screen "10_Startscreen" 800x480, template "01_Navigation"
   on GenerateScreen: SetTag("MainNavigationState", 1)
   GraphicView "Graphic view_2" at 0,0 size 800x480; Picture "PopUpBackground"
      Visibility <- "PopUpBackground"
   Button "Button_7" at 14,136 size 30x30; TextOff 'Text'
      Visibility <- "DB_HMI_Global_selection"
   Button "Button_10" at 14,195 size 30x30; TextOff 'Text'
      Visibility <- "DB_HMI_Global_selection"
   Button "Button_11" at 14,250 size 30x30; TextOff 'Text'
      Visibility <- "DB_HMI_Global_selection"
   Button "Button_13" at 14,311 size 30x30; TextOff 'Text'
      Visibility <- "DB_HMI_Global_selection"
   TextField "txtContentboard1" at 667,136 size 59x34; Text 'Calc. Time [s] / Name Parameter'
   TextField "txtContentboard1_1" at 723,141 size 65x24; Text 'Meas. Time [s] / Name Parameter'
   Button "Button_1" at 14,136 size 30x30; TextOff 'Text'
      on Click: SetTag("DB_HMI_Global_selection", 3)
   Button "Button_2" at 14,195 size 30x30; TextOff 'Text'
      on Click: SetTag("DB_HMI_Global_selection", 4)
   Button "Button_3" at 14,251 size 30x30; TextOff 'Text'
      on Click: SetTag("DB_HMI_Global_selection", 6)
   Button "Button_12" at 14,310 size 30x30; TextOff 'Text'
      on Click: SetTag("DB_HMI_Global_selection", 0)
   TextField "txtParameter1" at 82,159 size 99x24; Text 'Status / Parameter 1'
      Visibility <- "InScreenTabState"
   TextField "txtParameter1_1" at 82,199 size 99x24; Text 'Mode / Parameter 1'
      Visibility <- "InScreenTabState"
   TextField "txtParameter1_3" at 83,242 size 84x24; Text 'Producing car / Parameter 1'
      Visibility <- "InScreenTabState"
   TextField "Text field_4" at 32,381 size 142x20; Text 'Operation Commands'
   TextField "Text field_1" at 32,99 size 105x20; Text 'Production Line'
   TextField "txtParameter1_2" at 194,159 size 99x24; Text 'Status / Parameter 1'
      Visibility <- "InScreenTabState"
   TextField "txtParameter1_4" at 195,197 size 99x24; Text 'Mode / Parameter 1'
      Visibility <- "InScreenTabState"
   TextField "txtParameter1_5" at 195,242 size 84x24; Text 'Producing car / Parameter 1'
      Visibility <- "InScreenTabState"
   TextField "txtParameter1_6" at 306,159 size 99x24; Text 'Status / Parameter 1'
      Visibility <- "InScreenTabState"
   TextField "txtParameter1_7" at 307,197 size 99x24; Text 'Mode / Parameter 1'
      Visibility <- "InScreenTabState"
   TextField "txtParameter1_8" at 307,242 size 84x24; Text 'Producing car / Parameter 1'
      Visibility <- "InScreenTabState"
   TextField "txtParameter1_9" at 418,159 size 99x24; Text 'Status / Parameter 1'
      Visibility <- "InScreenTabState"
   TextField "txtParameter1_10" at 419,197 size 99x24; Text 'Mode / Parameter 1'
      Visibility <- "InScreenTabState"
   TextField "txtParameter1_11" at 419,242 size 84x24; Text 'Producing car / Parameter 1'
      Visibility <- "InScreenTabState"
   TextField "txtParameter1_12" at 530,159 size 99x24; Text 'Status / Parameter 1'
      Visibility <- "InScreenTabState"
   TextField "txtParameter1_13" at 531,197 size 99x24; Text 'Mode / Parameter 1'
      Visibility <- "InScreenTabState"
   TextField "txtParameter1_14" at 531,242 size 84x24; Text 'Producing car / Parameter 1'
      Visibility <- "InScreenTabState"
   GraphicView "Graphic view_1" at 46,139 size 25x25; Picture "Car_Red"
   GraphicView "Graphic view_3" at 47,196 size 25x25; Picture "Car_Green"
   GraphicView "Graphic view_4" at 47,251 size 25x25; Picture "Car_Blue_1"
   IOField "I/O field_1" at 671,168 size 56x24; FormatPattern 999
      ProcessValue <- "DB_HMI_ARG1_Seq1_Calculated_PT_Red(4)"
   TextField "txtTitleBar" at 80,128 size 55x24; Text 'Station 1 / Applikation'
   GraphicView "Graphic view_5" at 636,169 size 25x25; Picture "Car_Red"
   GraphicView "Graphic view_6" at 636,226 size 25x25; Picture "Car_Green"
   GraphicView "Graphic view_7" at 636,285 size 25x25; Picture "Car_Blue_1"
   TextField "txtTitleBar_1" at 200,122 size 55x24; Text 'Station 2 / Applikation'
   TextField "txtTitleBar_2" at 320,122 size 55x24; Text 'Station 3 / Applikation'
   TextField "txtTitleBar_3" at 440,122 size 55x24; Text 'Station 4 / Applikation'
   TextField "txtTitleBar_4" at 560,122 size 55x24; Text 'Station 5 / Applikation'
   Button "btnStart" at 184,377 size 119x29; TextOn 'STOP'; TextOff 'START'
      on Press: SetTag("DB_HMI_Global_Cmd_Start", 1); SetTag("DB_HMI_Global_Cmd_Start(1)", 1); SetTag("DB_HMI_Global_Cmd_Start(2)", 1); SetTag("DB_HMI_Global_Cmd_Start(3)", 1); SetTag("DB_HMI_Global_Cmd_Start(4)", 1)
      on Release: SetTag("DB_HMI_Global_Cmd_Start", 0); SetTag("DB_HMI_Global_Cmd_Start(1)", 0); SetTag("DB_HMI_Global_Cmd_Start(2)", 0); SetTag("DB_HMI_Global_Cmd_Start(3)", 0); SetTag("DB_HMI_Global_Cmd_Start(4)", 0)
   Button "btnStart_1" at 312,376 size 120x30; TextOn 'STOP'; TextOff 'STOP / START'
      on Release: SetTag("DB_HMI_Global_Cmd_Stop", 0); SetTag("DB_HMI_Global_Cmd_Stop(1)", 0); SetTag("DB_HMI_Global_Cmd_Stop(2)", 0); SetTag("DB_HMI_Global_Cmd_Stop(3)", 0); SetTag("DB_HMI_Global_Cmd_Stop(4)", 0)
      on Press: SetTag("DB_HMI_Global_Cmd_Stop", 1); SetTag("DB_HMI_Global_Cmd_Stop(1)", 1); SetTag("DB_HMI_Global_Cmd_Stop(2)", 1); SetTag("DB_HMI_Global_Cmd_Stop(3)", 1); SetTag("DB_HMI_Global_Cmd_Stop(4)", 1)
   IOField "I/O field_2" at 727,168 size 56x24; FormatPattern 999
      ProcessValue <- "DB_HMI_ARG1_Seq1_Messured_PT_Red(4)"
   TextField "txtTitleBar_5" at 192,128 size 55x24; Text 'Station 2 / Applikation'
   TextField "txtTitleBar_6" at 304,128 size 55x24; Text 'Station 3 / Applikation'
   TextField "txtTitleBar_7" at 416,128 size 55x24; Text 'Station 4 / Applikation'
   TextField "Text field_52" at 81,297 size 549x14; Text 'Text'
   TextField "txtTitleBar_8" at 528,128 size 55x24; Text 'Station 5 / Applikation'
   IOField "I/O field_3" at 671,224 size 56x24; FormatPattern 999
      ProcessValue <- "DB_HMI_ARG1_Seq1_Calculated_PT_Green(4)"
   IOField "I/O field_4" at 727,224 size 56x24; FormatPattern 999
      ProcessValue <- "DB_HMI_ARG1_Seq1_Messured_PT_Green(4)"
   IOField "I/O field_5" at 671,280 size 56x24; FormatPattern 999
      ProcessValue <- "DB_HMI_ARG1_Seq1_Calculated_PT_Blue(4)"
   IOField "I/O field_6" at 727,280 size 56x24; FormatPattern 999
      ProcessValue <- "DB_HMI_ARG1_Seq1_Messured_PT_Blue(4)"
   GraphicView "Grafikanzeige_1" at 46,312 size 26x22; Picture "Grafik_4"
   Button "btnState" at 143,133 size 39x25; TextOff '...'; PictureOff "More_Icon"
      on Click: ActivateScreen("21_Station_1", 0); SetTag("SubNavigationState", 2)
   Button "btnState_1" at 255,133 size 39x25; TextOff '...'; PictureOff "More_Icon"
      on Click: ActivateScreen("22_Station_2", 0); SetTag("SubNavigationState", 3)
   Button "btnState_2" at 367,133 size 39x25; TextOff '...'; PictureOff "More_Icon"
      on Click: ActivateScreen("23_Station_3", 0); SetTag("SubNavigationState", 4)
   Button "btnState_3" at 479,133 size 39x25; TextOff '...'; PictureOff "More_Icon"
      on Click: ActivateScreen("24_Station_4", 0); SetTag("SubNavigationState", 5)
   Button "btnState_4" at 591,133 size 39x25; TextOff '...'; PictureOff "More_Icon"
      on Click: ActivateScreen("25_Station_5", 0); SetTag("SubNavigationState", 6)
   Rectangle "rectState" at 0,48 size 56x38
      Appearance <- "CurrentMachineState"
   Button "btnState_5" at 201,53 size 34x31; TextOff '...'; PictureOff "More_Icon"
      on Click: ActivateScreen("11_Mode_Global", 0)
   TextField "Auto" at 67,63 size 35x20; Text 'Auto'
      Visibility <- "DB_HMI_Global_Status_Auto"
   TextField "Manual" at 69,63 size 34x20; Text 'Man'
      Visibility <- "DB_HMI_Global_Status_Man"
   TextField "txtStateHeadline" at 65,48 size 123x23; Text 'Mode / Status'
   Button "sTATUS" at 80,184 size 102x25; TextOff 'Text'; TextList "MachineStatus"
      on Activate: "VBFunction_1"()
      ProcessValue <- "status"
   Button "sTATUS_1" at 192,184 size 102x25; TextOff 'Text'; TextList "MachineStatus"
      ProcessValue <- "DB_HMI_ARG1_Seq1_Status_Busy(1)"
   Button "sTATUS_2" at 304,184 size 102x25; TextOff 'Text'; TextList "MachineStatus"
      ProcessValue <- "DB_HMI_ARG1_Seq1_Status_Busy(2)"
   Button "sTATUS_3" at 416,184 size 102x25; TextOff 'Text'; TextList "MachineStatus"
      ProcessValue <- "DB_HMI_ARG1_Seq1_Status_Busy(3)"
   Button "sTATUS_4" at 528,184 size 102x25; TextOff 'Text'; TextList "MachineStatus"
      ProcessValue <- "DB_HMI_ARG1_Seq1_Status_Busy(4)"
   Button "sTATUS_5" at 82,214 size 102x25; TextOff 'Text'; TextList "MachineMode"
      ProcessValue <- "DB_HMI_ARG1_Seq1_Status_Auto"
   Button "sTATUS_6" at 192,214 size 102x25; TextOff 'Text'; TextList "MachineMode"
      ProcessValue <- "DB_HMI_ARG1_Seq1_Status_Auto(1)"
   Button "sTATUS_7" at 304,214 size 102x25; TextOff 'Text'; TextList "MachineMode"
      ProcessValue <- "DB_HMI_ARG1_Seq1_Status_Auto(2)"
   Button "sTATUS_8" at 416,214 size 102x25; TextOff 'Text'; TextList "MachineMode"
      ProcessValue <- "DB_HMI_ARG1_Seq1_Status_Auto(3)"
   Button "sTATUS_9" at 528,214 size 102x25; TextOff 'Text'; TextList "MachineMode"
      ProcessValue <- "DB_HMI_ARG1_Seq1_Status_Auto(4)"
   Button "Button_4" at 101,274 size 60x60; TextOff 'Text'; PictureList "CarColorsGraph"
      ProcessValue <- "DB_HMI_inProduction"
   Button "Button_5" at 214,274 size 60x60; TextOff 'Text'; PictureList "CarColorsGraph"
      ProcessValue <- "DB_HMI_inProduction(1)"
   Button "Button_6" at 327,274 size 60x60; TextOff 'Text'; PictureList "CarColorsGraph"
      ProcessValue <- "DB_HMI_inProduction(2)"
   Button "Button_8" at 439,274 size 60x60; TextOff 'Text'; PictureList "CarColorsGraph"
      ProcessValue <- "DB_HMI_inProduction(3)"
   Button "Button_9" at 550,274 size 60x60; TextOff 'Text'; PictureList "CarColorsGraph"
      ProcessValue <- "DB_HMI_inProduction(4)"

screen "11_Mode_Global" 800x480
   Button "Button_5" at 299,208 size 88x48; TextOff 'Stop / AUTO'
      on Press: SetTag("DB_HMI_Global_Cmd_Auto", 1); SetTag("DB_HMI_Global_Cmd_Auto(1)", 1); SetTag("DB_HMI_Global_Cmd_Auto(2)", 1); SetTag("DB_HMI_Global_Cmd_Auto(3)", 1); SetTag("DB_HMI_Global_Cmd_Auto(4)", 1)
      on Release: SetTag("DB_HMI_Global_Cmd_Auto", 0); SetTag("DB_HMI_Global_Cmd_Auto(1)", 0); SetTag("DB_HMI_Global_Cmd_Auto(2)", 0); SetTag("DB_HMI_Global_Cmd_Auto(3)", 0); SetTag("DB_HMI_Global_Cmd_Auto(4)", 0)
   Button "Button_6" at 405,208 size 88x48; TextOff 'Reset / MAN'
      on Press: SetTag("DB_HMI_Global_Cmd_Man", 1); SetTag("DB_HMI_Global_Cmd_Man(1)", 1); SetTag("DB_HMI_Global_Cmd_Man(2)", 1); SetTag("DB_HMI_Global_Cmd_Man(3)", 1); SetTag("DB_HMI_Global_Cmd_Man(4)", 1)
      on Release: SetTag("DB_HMI_Global_Cmd_Man", 0); SetTag("DB_HMI_Global_Cmd_Man(1)", 0); SetTag("DB_HMI_Global_Cmd_Man(2)", 0); SetTag("DB_HMI_Global_Cmd_Man(3)", 0); SetTag("DB_HMI_Global_Cmd_Man(4)", 0)
   Button "Button_1" at 177,283 size 440x40; TextOn 'CLOSE / SCHLIESSEN'; TextOff 'CLOSE / SCHLIESSEN'
      on Click: function_efd93a16()
      Appearance <- "ButtonDown"
   TextField "txtTitleBar" at 16,8 size 495x32; Text 'Operating Mode / Betriebsmodus'
   TextField "txtParameter7_3" at 193,122 size 163x24; Text 'Current Mode / Aktueller Modus'
   TextField "Manual" at 193,148 size 35x20; Text 'Man'
      Visibility <- "DB_HMI_Global_Status_Man"
   TextField "Auto" at 193,149 size 41x20; Text 'Auto'
      Visibility <- "DB_HMI_Global_Status_Auto"

screen "21_Station_1" 800x480, template "01_Navigation"
   Button "Button_11" at 24,220 size 272x40; TextOff 'Simulate Values / Alle Quittieren'; PictureOff "More_Icon"
      on ReleaseLeft: ResetBit("Ext_AckSafety_DB_ack")
      on PressLeft: SetBit("Ext_AckSafety_DB_ack")
      on Click: ActivateScreen("40_SimValues_1", 0)
      on Press: ActivateScreen("40_SimValues_1", 0)
   Button "Button_1" at 24,324 size 272x40; TextOff 'Start / Alle Quittieren'; PictureOff "More_Icon"
      on Release: SetTag("DB_HMI_ARG1_Seq1_Cmd_Start", 0)
      on PressLeft: SetBit("Ext_AckSafety_DB_ack")
      on ReleaseLeft: ResetBit("Ext_AckSafety_DB_ack")
      on Press: SetTag("DB_HMI_ARG1_Seq1_Cmd_Start", 1); SetTag("DB_HMI_ARG1_Seq1_Cmd_Stop", 0)
      Visibility <- "DB_HMI_ARG1_Seq1_Status_Man"
      ObjectEnable <- "DB_HMI_ARG1_Seq1_Cmd_Start"
   Button "Button_2" at 24,376 size 272x40; TextOff 'Stop + Reset / Alle Quittieren'; PictureOff "More_Icon"
      on Release: SetTag("DB_HMI_ARG1_Seq1_Cmd_Stop", 0)
      on PressLeft: SetBit("Ext_AckSafety_DB_ack")
      on ReleaseLeft: ResetBit("Ext_AckSafety_DB_ack")
      on Press: SetTag("DB_HMI_ARG1_Seq1_Cmd_Stop", 1); SetTag("DB_HMI_ARG1_Seq1_Cmd_Start", 0)
      Visibility <- "DB_HMI_ARG1_Seq1_Status_Man"
      ObjectEnable <- "DB_HMI_ARG1_Seq1_Cmd_Stop"
   TextField "Text field_1" at 16,192 size 166x25; Text 'Simulation timers'
   TextField "Text field_2" at 16,296 size 105x25; Text 'Commands'
   TextField "Text field_26" at 564,176 size 204x24; Text 'Branch2'
   TextField "Text field_3" at 16,104 size 61x25; Text 'Status'
   TextField "Text field_16" at 344,176 size 204x24; Text 'Branch1'
   TextField "Text field_17" at 344,104 size 230x25; Text 'Running step sequences'
   Button "Button_3" at 218,123 size 45x45; TextOff 'Text'; PictureList "CarColorsGraph"
      Visibility <- "DB_HMI_ARG1_Seq1_Status_Auto"
      ProcessValue <- "DB_HMI_inProduction"
   TextField "Text field_4" at 180,104 size 118x27; Text 'Produced car'
   TextField "Text field_7" at 344,200 size 204x24; Text 'Step 1'
   TextField "Text field_5" at 344,224 size 204x24; Text 'Step 2'
   TextField "Text field_6" at 344,248 size 204x24; Text 'Step 3'
   TextField "Text field_8" at 344,272 size 204x24; Text 'Step 4'
   TextField "Text field_9" at 344,296 size 204x24; Text 'Step 5'
   TextField "Text field_10" at 344,320 size 204x24; Text 'Step 6'
   TextField "Text field_11" at 344,344 size 204x24; Text 'Step 7'
   TextField "Text field_12" at 344,368 size 204x24; Text 'Step 8'
   TextField "Text field_15" at 564,200 size 204x24; Text 'Step 1'
   TextField "Text field_18" at 564,224 size 204x24; Text 'Step 2'
   TextField "Text field_19" at 564,248 size 204x24; Text 'Step 3'
   TextField "Text field_20" at 564,272 size 204x24; Text 'Step 4'
   TextField "Text field_21" at 564,296 size 204x24; Text 'Step 5'
   TextField "Text field_22" at 564,320 size 204x24; Text 'Step 6'
   TextField "Text field_23" at 564,344 size 204x24; Text 'Step 7'
   TextField "Text field_24" at 564,368 size 204x24; Text 'Step 8'
   TextField "Text field_25" at 564,392 size 204x24; Text 'Step 9'
   TextField "Text field_13" at 344,392 size 204x24; Text 'Step 9'
   TextField "Text field_14" at 344,138 size 204x24; Text 'Step 0'
   TextField "Text field_52" at 344,200 size 204x24; Text 'Step 1'
      Visibility <- "DB_HMI_ARG1_Seq1_S2"
   TextField "Text field_27" at 344,224 size 204x24; Text 'Step 2'
      Visibility <- "DB_HMI_ARG1_Seq1_S3"
   TextField "Text field_28" at 344,249 size 204x24; Text 'Step 3'
      Visibility <- "DB_HMI_ARG1_Seq1_S4"
   TextField "Text field_29" at 344,272 size 204x24; Text 'Step 4'
      Visibility <- "DB_HMI_ARG1_Seq1_S5"
   TextField "Text field_30" at 344,296 size 204x24; Text 'Step 5'
      Visibility <- "DB_HMI_ARG1_Seq1_S6"
   TextField "Text field_31" at 344,320 size 204x24; Text 'Step 6'
      Visibility <- "DB_HMI_ARG1_Seq1_S7"
   TextField "Text field_32" at 344,344 size 204x24; Text 'Step 7'
      Visibility <- "DB_HMI_ARG1_Seq1_S8"
   TextField "Text field_33" at 344,368 size 204x24; Text 'Step 8'
      Visibility <- "DB_HMI_ARG1_Seq1_S9"
   TextField "Text field_34" at 344,392 size 204x24; Text 'Step 9'
      Visibility <- "DB_HMI_ARG1_Seq1_S10"
   TextField "Text field_35" at 564,200 size 204x24; Text 'Step 1'
      Visibility <- "DB_HMI_ARG1_Seq1_S11"
   TextField "Text field_36" at 564,224 size 204x24; Text 'Step 2'
      Visibility <- "DB_HMI_ARG1_Seq1_S12"
   TextField "Text field_37" at 564,248 size 204x24; Text 'Step 3'
      Visibility <- "DB_HMI_ARG1_Seq1_S13"
   TextField "Text field_38" at 564,272 size 204x24; Text 'Step 4'
      Visibility <- "DB_HMI_ARG1_Seq1_S14"
   TextField "Text field_39" at 564,296 size 204x24; Text 'Step 5'
      Visibility <- "DB_HMI_ARG1_Seq1_S15"
   TextField "Text field_40" at 564,320 size 204x24; Text 'Step 6'
      Visibility <- "DB_HMI_ARG1_Seq1_S16"
   TextField "Text field_41" at 564,344 size 204x24; Text 'Step 7'
      Visibility <- "DB_HMI_ARG1_Seq1_S17"
   TextField "Text field_42" at 564,368 size 204x24; Text 'Step 8'
      Visibility <- "DB_HMI_ARG1_Seq1_S18"
   TextField "Text field_43" at 564,392 size 204x24; Text 'Step 9'
      Visibility <- "DB_HMI_ARG1_Seq1_S19"
   TextField "Text field_44" at 344,138 size 204x24; Text 'Step 0'
      Visibility <- "DB_HMI_ARG1_Seq1_S1"
   SymbolicIOField "Symbolic I/O field_1" at 182,129 size 117x32; TextOn '1'; TextOff '0'; TextList "Car_color"
      ProcessValue <- "DB_HMI_dropdown_selection"
      Visibility <- "DB_HMI_ARG1_Seq1_Status_Man"
   TextField "Busy" at 14,134 size 41x22; Text 'Busy'
      Visibility <- "DB_HMI_ARG1_Seq1_Status_Busy"
   TextField "Idle" at 14,134 size 35x22; Text 'Idle'
      Visibility <- "DB_HMI_ARG1_Seq1_Status_Idle"
   Rectangle "rectState" at 0,48 size 56x38
      Appearance <- "CurrentMachineState"
   Button "btnState" at 201,53 size 34x31; TextOff '...'; PictureOff "More_Icon"
      on Click: ActivateScreen("31_Mode_Station_1", 0)
   TextField "Auto" at 67,63 size 35x20; Text 'Auto'
      Visibility <- "DB_HMI_ARG1_Seq1_Status_Auto"
   TextField "Manual" at 69,63 size 34x20; Text 'Man'
      Visibility <- "DB_HMI_ARG1_Seq1_Status_Man"
   TextField "txtStateHeadline" at 65,48 size 123x23; Text 'Mode / Status'

screen "22_Station_2" 800x480, template "01_Navigation"
   Button "Button_11" at 24,220 size 272x40; TextOff 'Simulate Values / Alle Quittieren'; PictureOff "More_Icon"
      on ReleaseLeft: ResetBit("Ext_AckSafety_DB_ack")
      on PressLeft: SetBit("Ext_AckSafety_DB_ack")
      on Click: ActivateScreen("40_SimValues_2", 0)
   Button "Button_1" at 24,324 size 272x40; TextOff 'Start / Alle Quittieren'; PictureOff "More_Icon"
      on Release: SetTag("DB_HMI_ARG1_Seq1_Cmd_Start(1)", 0)
      on PressLeft: SetBit("Ext_AckSafety_DB_ack")
      on ReleaseLeft: ResetBit("Ext_AckSafety_DB_ack")
      on Press: SetTag("DB_HMI_ARG1_Seq1_Cmd_Start(1)", 1); SetTag("DB_HMI_ARG1_Seq1_Cmd_Stop(1)", 0)
      Visibility <- "DB_HMI_ARG1_Seq1_Status_Man(1)"
      ObjectEnable <- "DB_HMI_ARG1_Seq1_Cmd_Start(1)"
   Button "Button_2" at 24,376 size 272x40; TextOff 'Stop + Reset / Alle Quittieren'; PictureOff "More_Icon"
      on Release: SetTag("DB_HMI_ARG1_Seq1_Cmd_Stop(1)", 0)
      on PressLeft: SetBit("Ext_AckSafety_DB_ack")
      on ReleaseLeft: ResetBit("Ext_AckSafety_DB_ack")
      on Press: SetTag("DB_HMI_ARG1_Seq1_Cmd_Stop(1)", 1); SetTag("DB_HMI_ARG1_Seq1_Cmd_Start(1)", 0)
      Visibility <- "DB_HMI_ARG1_Seq1_Status_Man(1)"
      ObjectEnable <- "DB_HMI_ARG1_Seq1_Cmd_Stop(1)"
   TextField "Text field_1" at 16,192 size 166x25; Text 'Simulation timers'
   TextField "Text field_2" at 16,296 size 105x25; Text 'Commands'
   TextField "Text field_26" at 564,176 size 204x24; Text 'Branch2'
   TextField "Text field_3" at 16,104 size 61x25; Text 'Status'
   TextField "Text field_16" at 344,176 size 204x24; Text 'Branch1'
   SymbolicIOField "DropDownCars" at 182,129 size 117x32; TextOn '1'; TextOff '0'; TextList "Car_color"
      ProcessValue <- "DB_HMI_dropdown_selection(1)"
      Visibility <- "DB_HMI_ARG1_Seq1_Status_Man(1)"
   TextField "Text field_17" at 344,104 size 230x25; Text 'Running step sequences'
   TextField "Text field_4" at 180,104 size 118x27; Text 'Produced car'
   Button "Button_3" at 218,123 size 45x45; TextOff 'Text'; PictureList "CarColorsGraph"
      Visibility <- "DB_HMI_ARG1_Seq1_Status_Auto(1)"
      ProcessValue <- "DB_HMI_inProduction(1)"
   TextField "Text field_7" at 344,200 size 204x24; Text 'Step 1'
   TextField "Text field_5" at 344,224 size 204x24; Text 'Step 2'
   TextField "Text field_6" at 344,248 size 204x24; Text 'Step 3'
   TextField "Text field_8" at 344,272 size 204x24; Text 'Step 4'
   TextField "Text field_9" at 344,296 size 204x24; Text 'Step 5'
   TextField "Text field_10" at 344,320 size 204x24; Text 'Step 6'
   TextField "Text field_11" at 344,344 size 204x24; Text 'Step 7'
   TextField "Text field_12" at 344,368 size 204x24; Text 'Step 8'
   TextField "Text field_15" at 564,200 size 204x24; Text 'Step 1'
   TextField "Text field_18" at 564,224 size 204x24; Text 'Step 2'
   TextField "Text field_19" at 564,248 size 204x24; Text 'Step 3'
   TextField "Text field_20" at 564,272 size 204x24; Text 'Step 4'
   TextField "Text field_21" at 564,296 size 204x24; Text 'Step 5'
   TextField "Text field_22" at 564,320 size 204x24; Text 'Step 6'
   TextField "Text field_23" at 564,344 size 204x24; Text 'Step 7'
   TextField "Text field_24" at 564,368 size 204x24; Text 'Step 8'
   TextField "Text field_25" at 564,392 size 204x24; Text 'Step 9'
   TextField "Text field_13" at 344,392 size 204x24; Text 'Step 9'
   TextField "Text field_14" at 344,138 size 204x24; Text 'Step 0'
   TextField "Text field_52" at 344,200 size 204x24; Text 'Step 1'
      Visibility <- "DB_HMI_ARG1_Seq1_S2(1)"
   TextField "Text field_27" at 344,224 size 204x24; Text 'Step 2'
      Visibility <- "DB_HMI_ARG1_Seq1_S3(1)"
   TextField "Text field_28" at 344,249 size 204x24; Text 'Step 3'
      Visibility <- "DB_HMI_ARG1_Seq1_S4(1)"
   TextField "Text field_29" at 344,272 size 204x24; Text 'Step 4'
      Visibility <- "DB_HMI_ARG1_Seq1_S5(1)"
   TextField "Text field_30" at 344,296 size 204x24; Text 'Step 5'
      Visibility <- "DB_HMI_ARG1_Seq1_S6(1)"
   TextField "Text field_31" at 344,320 size 204x24; Text 'Step 6'
      Visibility <- "DB_HMI_ARG1_Seq1_S7(1)"
   TextField "Text field_32" at 344,344 size 204x24; Text 'Step 7'
      Visibility <- "DB_HMI_ARG1_Seq1_S8(1)"
   TextField "Text field_33" at 344,368 size 204x24; Text 'Step 8'
      Visibility <- "DB_HMI_ARG1_Seq1_S9(1)"
   TextField "Text field_34" at 344,392 size 204x24; Text 'Step 9'
      Visibility <- "DB_HMI_ARG1_Seq1_S10(1)"
   TextField "Text field_35" at 564,200 size 204x24; Text 'Step 1'
      Visibility <- "DB_HMI_ARG1_Seq1_S11(1)"
   TextField "Text field_36" at 564,224 size 204x24; Text 'Step 2'
      Visibility <- "DB_HMI_ARG1_Seq1_S12(1)"
   TextField "Text field_37" at 564,248 size 204x24; Text 'Step 3'
      Visibility <- "DB_HMI_ARG1_Seq1_S13(1)"
   TextField "Text field_38" at 564,272 size 204x24; Text 'Step 4'
      Visibility <- "DB_HMI_ARG1_Seq1_S14(1)"
   TextField "Text field_39" at 564,296 size 204x24; Text 'Step 5'
      Visibility <- "DB_HMI_ARG1_Seq1_S15(1)"
   TextField "Text field_40" at 564,320 size 204x24; Text 'Step 6'
      Visibility <- "DB_HMI_ARG1_Seq1_S16(1)"
   TextField "Text field_41" at 564,344 size 204x24; Text 'Step 7'
      Visibility <- "DB_HMI_ARG1_Seq1_S17(1)"
   TextField "Text field_42" at 564,368 size 204x24; Text 'Step 8'
      Visibility <- "DB_HMI_ARG1_Seq1_S18(1)"
   TextField "Text field_43" at 564,392 size 204x24; Text 'Step 9'
      Visibility <- "DB_HMI_ARG1_Seq1_S19(1)"
   TextField "Text field_44" at 344,138 size 204x24; Text 'Step 0'
      Visibility <- "DB_HMI_ARG1_Seq1_S1(1)"
   TextField "Busy" at 14,134 size 41x22; Text 'Busy'
      Visibility <- "DB_HMI_ARG1_Seq1_Status_Busy(1)"
   TextField "Idle" at 14,134 size 35x22; Text 'Idle'
      Visibility <- "DB_HMI_ARG1_Seq1_Status_Idle(1)"
   Rectangle "rectState" at 0,48 size 56x38
      Appearance <- "CurrentMachineState"
   Button "btnState" at 201,53 size 34x31; TextOff '...'; PictureOff "More_Icon"
      on Click: ActivateScreen("32_Mode_Station_2", 0)
   TextField "Auto" at 67,63 size 35x20; Text 'Auto'
      Visibility <- "DB_HMI_ARG1_Seq1_Status_Auto(1)"
   TextField "Manual" at 69,63 size 34x20; Text 'Man'
      Visibility <- "DB_HMI_ARG1_Seq1_Status_Man(1)"
   TextField "txtStateHeadline" at 65,48 size 123x23; Text 'Mode / Status'

screen "23_Station_3" 800x480, template "01_Navigation"
   Button "Button_11" at 24,220 size 272x40; TextOff 'Simulate Values / Alle Quittieren'; PictureOff "More_Icon"
      on ReleaseLeft: ResetBit("Ext_AckSafety_DB_ack")
      on PressLeft: SetBit("Ext_AckSafety_DB_ack")
      on Click: ActivateScreen("40_SimValues_3", 0)
   Button "Button_1" at 24,324 size 272x40; TextOff 'Start / Alle Quittieren'; PictureOff "More_Icon"
      on Release: SetTag("DB_HMI_ARG1_Seq1_Cmd_Start(2)", 0)
      on PressLeft: SetBit("Ext_AckSafety_DB_ack")
      on ReleaseLeft: ResetBit("Ext_AckSafety_DB_ack")
      on Press: SetTag("DB_HMI_ARG1_Seq1_Cmd_Start(2)", 1); SetTag("DB_HMI_ARG1_Seq1_Cmd_Stop(2)", 0)
      ObjectEnable <- "DB_HMI_ARG1_Seq1_Cmd_Start"
      Visibility <- "DB_HMI_ARG1_Seq1_Status_Man(2)"
   Button "Button_2" at 24,376 size 272x40; TextOff 'Stop + Reset / Alle Quittieren'; PictureOff "More_Icon"
      on Release: SetTag("DB_HMI_ARG1_Seq1_Cmd_Stop(2)", 0)
      on PressLeft: SetBit("Ext_AckSafety_DB_ack")
      on ReleaseLeft: ResetBit("Ext_AckSafety_DB_ack")
      on Press: SetTag("DB_HMI_ARG1_Seq1_Cmd_Stop(2)", 1)
      ObjectEnable <- "DB_HMI_ARG1_Seq1_Cmd_Stop"
      Visibility <- "DB_HMI_ARG1_Seq1_Status_Man(2)"
   TextField "Text field_1" at 16,192 size 166x25; Text 'Simulation timers'
   TextField "Text field_2" at 16,296 size 105x25; Text 'Commands'
   TextField "Text field_26" at 564,176 size 204x24; Text 'Branch2'
   TextField "Text field_3" at 16,104 size 61x25; Text 'Status'
   TextField "Text field_16" at 344,176 size 204x24; Text 'Branch1'
   SymbolicIOField "DropDownCars" at 182,129 size 117x32; TextOn '1'; TextOff '0'; TextList "Car_color"
      ProcessValue <- "DB_HMI_dropdown_selection(2)"
      Visibility <- "DB_HMI_ARG1_Seq1_Status_Man(2)"
   TextField "Text field_17" at 344,104 size 230x25; Text 'Running step sequences'
   TextField "Text field_4" at 180,104 size 118x27; Text 'Produced car'
   Button "Button_3" at 218,123 size 45x45; TextOff 'Text'; PictureList "CarColorsGraph"
      Visibility <- "DB_HMI_ARG1_Seq1_Status_Auto(2)"
      ProcessValue <- "DB_HMI_inProduction(2)"
   TextField "Text field_7" at 344,200 size 204x24; Text 'Step 1'
   TextField "Text field_5" at 344,224 size 204x24; Text 'Step 2'
   TextField "Text field_6" at 344,248 size 204x24; Text 'Step 3'
   TextField "Text field_8" at 344,272 size 204x24; Text 'Step 4'
   TextField "Text field_9" at 344,296 size 204x24; Text 'Step 5'
   TextField "Text field_10" at 344,320 size 204x24; Text 'Step 6'
   TextField "Text field_11" at 344,344 size 204x24; Text 'Step 7'
   TextField "Text field_12" at 344,368 size 204x24; Text 'Step 8'
   TextField "Text field_15" at 564,200 size 204x24; Text 'Step 1'
   TextField "Text field_18" at 564,224 size 204x24; Text 'Step 2'
   TextField "Text field_19" at 564,248 size 204x24; Text 'Step 3'
   TextField "Text field_20" at 564,272 size 204x24; Text 'Step 4'
   TextField "Text field_21" at 564,296 size 204x24; Text 'Step 5'
   TextField "Text field_22" at 564,320 size 204x24; Text 'Step 6'
   TextField "Text field_23" at 564,344 size 204x24; Text 'Step 7'
   TextField "Text field_24" at 564,368 size 204x24; Text 'Step 8'
   TextField "Text field_25" at 564,392 size 204x24; Text 'Step 9'
   TextField "Text field_13" at 344,392 size 204x24; Text 'Step 9'
   TextField "Text field_14" at 344,138 size 204x24; Text 'Step 0'
   TextField "Text field_52" at 344,200 size 204x24; Text 'Step 1'
      Visibility <- "DB_HMI_ARG1_Seq1_S2(2)"
   TextField "Text field_27" at 344,224 size 204x24; Text 'Step 2'
      Visibility <- "DB_HMI_ARG1_Seq1_S3(2)"
   TextField "Text field_28" at 344,249 size 204x24; Text 'Step 3'
      Visibility <- "DB_HMI_ARG1_Seq1_S4(2)"
   TextField "Text field_29" at 344,272 size 204x24; Text 'Step 4'
      Visibility <- "DB_HMI_ARG1_Seq1_S5(2)"
   TextField "Text field_30" at 344,296 size 204x24; Text 'Step 5'
      Visibility <- "DB_HMI_ARG1_Seq1_S6(2)"
   TextField "Text field_31" at 344,320 size 204x24; Text 'Step 6'
      Visibility <- "DB_HMI_ARG1_Seq1_S7(2)"
   TextField "Text field_32" at 344,344 size 204x24; Text 'Step 7'
      Visibility <- "DB_HMI_ARG1_Seq1_S8(2)"
   TextField "Text field_33" at 344,368 size 204x24; Text 'Step 8'
      Visibility <- "DB_HMI_ARG1_Seq1_S9(2)"
   TextField "Text field_34" at 344,392 size 204x24; Text 'Step 9'
      Visibility <- "DB_HMI_ARG1_Seq1_S10(2)"
   TextField "Text field_35" at 564,200 size 204x24; Text 'Step 1'
      Visibility <- "DB_HMI_ARG1_Seq1_S11(2)"
   TextField "Text field_36" at 564,224 size 204x24; Text 'Step 2'
      Visibility <- "DB_HMI_ARG1_Seq1_S12(2)"
   TextField "Text field_37" at 564,248 size 204x24; Text 'Step 3'
      Visibility <- "DB_HMI_ARG1_Seq1_S13(2)"
   TextField "Text field_38" at 564,272 size 204x24; Text 'Step 4'
      Visibility <- "DB_HMI_ARG1_Seq1_S14(2)"
   TextField "Text field_39" at 564,296 size 204x24; Text 'Step 5'
      Visibility <- "DB_HMI_ARG1_Seq1_S15(2)"
   TextField "Text field_40" at 564,320 size 204x24; Text 'Step 6'
      Visibility <- "DB_HMI_ARG1_Seq1_S16(2)"
   TextField "Text field_41" at 564,344 size 204x24; Text 'Step 7'
      Visibility <- "DB_HMI_ARG1_Seq1_S17(2)"
   TextField "Text field_42" at 564,368 size 204x24; Text 'Step 8'
      Visibility <- "DB_HMI_ARG1_Seq1_S18(2)"
   TextField "Text field_43" at 564,392 size 204x24; Text 'Step 9'
      Visibility <- "DB_HMI_ARG1_Seq1_S19(2)"
   TextField "Text field_44" at 344,138 size 204x24; Text 'Step 0'
      Visibility <- "DB_HMI_ARG1_Seq1_S1(2)"
   TextField "Busy" at 14,134 size 41x22; Text 'Busy'
      Visibility <- "DB_HMI_ARG1_Seq1_Status_Busy(2)"
   TextField "Idle" at 14,134 size 35x22; Text 'Idle'
      Visibility <- "DB_HMI_ARG1_Seq1_Status_Idle(2)"
   Rectangle "rectState" at 0,48 size 56x38
      Appearance <- "CurrentMachineState"
   Button "btnState" at 201,53 size 34x31; TextOff '...'; PictureOff "More_Icon"
      on Click: ActivateScreen("33_Mode_Station_3", 0)
   TextField "Auto" at 67,63 size 35x20; Text 'Auto'
      Visibility <- "DB_HMI_ARG1_Seq1_Status_Auto(2)"
   TextField "Manual" at 69,63 size 34x20; Text 'Man'
      Visibility <- "DB_HMI_ARG1_Seq1_Status_Man(2)"
   TextField "txtStateHeadline" at 65,48 size 123x23; Text 'Mode / Status'

screen "24_Station_4" 800x480, template "01_Navigation"
   Button "Button_11" at 24,220 size 272x40; TextOff 'Simulate Values / Alle Quittieren'; PictureOff "More_Icon"
      on ReleaseLeft: ResetBit("Ext_AckSafety_DB_ack")
      on PressLeft: SetBit("Ext_AckSafety_DB_ack")
      on Click: ActivateScreen("40_SimValues_4", 0)
   Button "Button_1" at 24,324 size 272x40; TextOff 'Start / Alle Quittieren'; PictureOff "More_Icon"
      on Release: SetTag("DB_HMI_ARG1_Seq1_Cmd_Start(3)", 0)
      on PressLeft: SetBit("Ext_AckSafety_DB_ack")
      on ReleaseLeft: ResetBit("Ext_AckSafety_DB_ack")
      on Press: SetTag("DB_HMI_ARG1_Seq1_Cmd_Start(3)", 1)
      ObjectEnable <- "DB_HMI_ARG1_Seq1_Cmd_Start"
      Visibility <- "DB_HMI_ARG1_Seq1_Status_Man(3)"
   Button "Button_2" at 24,376 size 272x40; TextOff 'Stop + Reset / Alle Quittieren'; PictureOff "More_Icon"
      on Release: SetTag("DB_HMI_ARG1_Seq1_Cmd_Stop(3)", 0)
      on PressLeft: SetBit("Ext_AckSafety_DB_ack")
      on ReleaseLeft: ResetBit("Ext_AckSafety_DB_ack")
      on Press: SetTag("DB_HMI_ARG1_Seq1_Cmd_Stop(3)", 1)
      ObjectEnable <- "DB_HMI_ARG1_Seq1_Cmd_Stop"
      Visibility <- "DB_HMI_ARG1_Seq1_Status_Man(3)"
   TextField "Text field_1" at 16,192 size 166x25; Text 'Simulation timers'
   TextField "Text field_2" at 16,296 size 105x25; Text 'Commands'
   TextField "Text field_26" at 564,176 size 204x24; Text 'Branch2'
   TextField "Text field_3" at 16,104 size 61x25; Text 'Status'
   TextField "Text field_16" at 344,176 size 204x24; Text 'Branch1'
   TextField "Text field_17" at 344,104 size 230x25; Text 'Running step sequences'
   TextField "Text field_4" at 180,104 size 118x27; Text 'Produced car'
   Button "Button_3" at 218,123 size 45x45; TextOff 'Text'; PictureList "CarColorsGraph"
      Visibility <- "DB_HMI_ARG1_Seq1_Status_Auto(3)"
      ProcessValue <- "DB_HMI_inProduction(3)"
   TextField "Text field_7" at 344,200 size 204x24; Text 'Step 1'
   TextField "Text field_5" at 344,224 size 204x24; Text 'Step 2'
   TextField "Text field_6" at 344,248 size 204x24; Text 'Step 3'
   TextField "Text field_8" at 344,272 size 204x24; Text 'Step 4'
   TextField "Text field_9" at 344,296 size 204x24; Text 'Step 5'
   TextField "Text field_10" at 344,320 size 204x24; Text 'Step 6'
   TextField "Text field_11" at 344,344 size 204x24; Text 'Step 7'
   TextField "Text field_12" at 344,368 size 204x24; Text 'Step 8'
   TextField "Text field_15" at 564,200 size 204x24; Text 'Step 1'
   TextField "Text field_18" at 564,224 size 204x24; Text 'Step 2'
   TextField "Text field_19" at 564,248 size 204x24; Text 'Step 3'
   TextField "Text field_20" at 564,272 size 204x24; Text 'Step 4'
   TextField "Text field_21" at 564,296 size 204x24; Text 'Step 5'
   TextField "Text field_22" at 564,320 size 204x24; Text 'Step 6'
   TextField "Text field_23" at 564,344 size 204x24; Text 'Step 7'
   TextField "Text field_24" at 564,368 size 204x24; Text 'Step 8'
   TextField "Text field_25" at 564,392 size 204x24; Text 'Step 9'
   TextField "Text field_13" at 344,392 size 204x24; Text 'Step 9'
   TextField "Text field_14" at 344,138 size 204x24; Text 'Step 0'
   TextField "Text field_52" at 344,200 size 204x24; Text 'Step 1'
      Visibility <- "DB_HMI_ARG1_Seq1_S2(3)"
   TextField "Text field_27" at 344,224 size 204x24; Text 'Step 2'
      Visibility <- "DB_HMI_ARG1_Seq1_S3(3)"
   TextField "Text field_28" at 344,249 size 204x24; Text 'Step 3'
      Visibility <- "DB_HMI_ARG1_Seq1_S4(3)"
   TextField "Text field_29" at 344,272 size 204x24; Text 'Step 4'
      Visibility <- "DB_HMI_ARG1_Seq1_S5(3)"
   TextField "Text field_30" at 344,296 size 204x24; Text 'Step 5'
      Visibility <- "DB_HMI_ARG1_Seq1_S6(3)"
   TextField "Text field_31" at 344,320 size 204x24; Text 'Step 6'
      Visibility <- "DB_HMI_ARG1_Seq1_S7(3)"
   TextField "Text field_32" at 344,344 size 204x24; Text 'Step 7'
      Visibility <- "DB_HMI_ARG1_Seq1_S8(3)"
   TextField "Text field_33" at 344,368 size 204x24; Text 'Step 8'
      Visibility <- "DB_HMI_ARG1_Seq1_S9(3)"
   TextField "Text field_34" at 344,392 size 204x24; Text 'Step 9'
      Visibility <- "DB_HMI_ARG1_Seq1_S10(3)"
   TextField "Text field_35" at 564,200 size 204x24; Text 'Step 1'
      Visibility <- "DB_HMI_ARG1_Seq1_S11(3)"
   TextField "Text field_36" at 564,224 size 204x24; Text 'Step 2'
      Visibility <- "DB_HMI_ARG1_Seq1_S12(3)"
   TextField "Text field_37" at 564,248 size 204x24; Text 'Step 3'
      Visibility <- "DB_HMI_ARG1_Seq1_S13(3)"
   TextField "Text field_38" at 564,272 size 204x24; Text 'Step 4'
      Visibility <- "DB_HMI_ARG1_Seq1_S14(3)"
   TextField "Text field_39" at 564,296 size 204x24; Text 'Step 5'
      Visibility <- "DB_HMI_ARG1_Seq1_S15(3)"
   TextField "Text field_40" at 564,320 size 204x24; Text 'Step 6'
      Visibility <- "DB_HMI_ARG1_Seq1_S16(3)"
   TextField "Text field_41" at 564,344 size 204x24; Text 'Step 7'
      Visibility <- "DB_HMI_ARG1_Seq1_S17(3)"
   TextField "Text field_42" at 564,368 size 204x24; Text 'Step 8'
      Visibility <- "DB_HMI_ARG1_Seq1_S18(3)"
   TextField "Text field_43" at 564,392 size 204x24; Text 'Step 9'
      Visibility <- "DB_HMI_ARG1_Seq1_S19(3)"
   TextField "Text field_44" at 344,138 size 204x24; Text 'Step 0'
      Visibility <- "DB_HMI_ARG1_Seq1_S1(3)"
   SymbolicIOField "DropDownCars" at 182,129 size 117x32; TextOn '1'; TextOff '0'; TextList "Car_color"
      ProcessValue <- "DB_HMI_dropdown_selection(3)"
      Visibility <- "DB_HMI_ARG1_Seq1_Status_Man(3)"
   TextField "Busy" at 14,134 size 41x22; Text 'Busy'
      Visibility <- "DB_HMI_ARG1_Seq1_Status_Busy(3)"
   TextField "Idle" at 14,134 size 35x22; Text 'Idle'
      Visibility <- "DB_HMI_ARG1_Seq1_Status_Idle(3)"
   Rectangle "rectState" at 0,48 size 56x38
      Appearance <- "CurrentMachineState"
   Button "btnState" at 201,53 size 34x31; TextOff '...'; PictureOff "More_Icon"
      on Click: ActivateScreen("34_Mode_Station_4", 0)
   TextField "Auto" at 67,63 size 35x20; Text 'Auto'
      Visibility <- "DB_HMI_ARG1_Seq1_Status_Auto(3)"
   TextField "Manual" at 69,63 size 34x20; Text 'Man'
      Visibility <- "DB_HMI_ARG1_Seq1_Status_Man(3)"
   TextField "txtStateHeadline" at 65,48 size 123x23; Text 'Mode / Status'

screen "25_Station_5" 800x480, template "01_Navigation"
   Button "Button_11" at 24,220 size 272x40; TextOff 'Simulate Values / Alle Quittieren'; PictureOff "More_Icon"
      on ReleaseLeft: ResetBit("Ext_AckSafety_DB_ack")
      on PressLeft: SetBit("Ext_AckSafety_DB_ack")
      on Click: ActivateScreen("40_SimValues_5", 0)
   Button "Button_1" at 24,324 size 272x40; TextOff 'Start / Alle Quittieren'; PictureOff "More_Icon"
      on Release: SetTag("DB_HMI_ARG1_Seq1_Cmd_Start(4)", 0)
      on PressLeft: SetBit("Ext_AckSafety_DB_ack")
      on ReleaseLeft: ResetBit("Ext_AckSafety_DB_ack")
      on Press: SetTag("DB_HMI_ARG1_Seq1_Cmd_Start(4)", 1)
      ObjectEnable <- "DB_HMI_ARG1_Seq1_Cmd_Start"
      Visibility <- "DB_HMI_ARG1_Seq1_Status_Man(4)"
   Button "Button_2" at 24,376 size 272x40; TextOff 'Stop + Reset / Alle Quittieren'; PictureOff "More_Icon"
      on Release: SetTag("DB_HMI_ARG1_Seq1_Cmd_Stop(4)", 0)
      on PressLeft: SetBit("Ext_AckSafety_DB_ack")
      on ReleaseLeft: ResetBit("Ext_AckSafety_DB_ack")
      on Press: SetTag("DB_HMI_ARG1_Seq1_Cmd_Stop(4)", 1)
      ObjectEnable <- "DB_HMI_ARG1_Seq1_Cmd_Stop"
      Visibility <- "DB_HMI_ARG1_Seq1_Status_Man(4)"
   TextField "Text field_1" at 16,192 size 166x25; Text 'Simulation timers'
   TextField "Text field_2" at 16,296 size 105x25; Text 'Commands'
   TextField "Text field_26" at 564,176 size 204x24; Text 'Branch2'
   TextField "Text field_3" at 16,104 size 61x25; Text 'Status'
   TextField "Text field_16" at 344,176 size 204x24; Text 'Branch1'
   SymbolicIOField "DropDownCars" at 182,129 size 117x32; TextOn '1'; TextOff '0'; TextList "Car_color"
      ProcessValue <- "DB_HMI_dropdown_selection(4)"
      Visibility <- "DB_HMI_ARG1_Seq1_Status_Man(4)"
   TextField "Text field_17" at 344,104 size 230x25; Text 'Running step sequences'
   TextField "Text field_4" at 180,104 size 118x27; Text 'Produced car'
   Button "Button_3" at 218,123 size 45x45; TextOff 'Text'; PictureList "CarColorsGraph"
      Visibility <- "DB_HMI_ARG1_Seq1_Status_Auto(4)"
      ProcessValue <- "DB_HMI_inProduction(4)"
   TextField "Text field_7" at 344,200 size 204x24; Text 'Step 1'
   TextField "Text field_5" at 344,224 size 204x24; Text 'Step 2'
   TextField "Text field_6" at 344,248 size 204x24; Text 'Step 3'
   TextField "Text field_8" at 344,272 size 204x24; Text 'Step 4'
   TextField "Text field_9" at 344,296 size 204x24; Text 'Step 5'
   TextField "Text field_10" at 344,320 size 204x24; Text 'Step 6'
   TextField "Text field_11" at 344,344 size 204x24; Text 'Step 7'
   TextField "Text field_12" at 344,368 size 204x24; Text 'Step 8'
   TextField "Text field_15" at 564,200 size 204x24; Text 'Step 1'
   TextField "Text field_18" at 564,224 size 204x24; Text 'Step 2'
   TextField "Text field_19" at 564,248 size 204x24; Text 'Step 3'
   TextField "Text field_20" at 564,272 size 204x24; Text 'Step 4'
   TextField "Text field_21" at 564,296 size 204x24; Text 'Step 5'
   TextField "Text field_22" at 564,320 size 204x24; Text 'Step 6'
   TextField "Text field_23" at 564,344 size 204x24; Text 'Step 7'
   TextField "Text field_24" at 564,368 size 204x24; Text 'Step 8'
   TextField "Text field_25" at 564,392 size 204x24; Text 'Step 9'
   TextField "Text field_13" at 344,392 size 204x24; Text 'Step 9'
   TextField "Text field_14" at 344,138 size 204x24; Text 'Step 0'
   TextField "Text field_52" at 344,200 size 204x24; Text 'Step 1'
      Visibility <- "DB_HMI_ARG1_Seq1_S2(4)"
   TextField "Text field_27" at 344,224 size 204x24; Text 'Step 2'
      Visibility <- "DB_HMI_ARG1_Seq1_S3(4)"
   TextField "Text field_28" at 344,249 size 204x24; Text 'Step 3'
      Visibility <- "DB_HMI_ARG1_Seq1_S4(4)"
   TextField "Text field_29" at 344,272 size 204x24; Text 'Step 4'
      Visibility <- "DB_HMI_ARG1_Seq1_S5(4)"
   TextField "Text field_30" at 344,296 size 204x24; Text 'Step 5'
      Visibility <- "DB_HMI_ARG1_Seq1_S6(4)"
   TextField "Text field_31" at 344,320 size 204x24; Text 'Step 6'
      Visibility <- "DB_HMI_ARG1_Seq1_S7(4)"
   TextField "Text field_32" at 344,344 size 204x24; Text 'Step 7'
      Visibility <- "DB_HMI_ARG1_Seq1_S8(4)"
   TextField "Text field_33" at 344,368 size 204x24; Text 'Step 8'
      Visibility <- "DB_HMI_ARG1_Seq1_S9(4)"
   TextField "Text field_34" at 344,392 size 204x24; Text 'Step 9'
      Visibility <- "DB_HMI_ARG1_Seq1_S10(4)"
   TextField "Text field_35" at 564,200 size 204x24; Text 'Step 1'
      Visibility <- "DB_HMI_ARG1_Seq1_S11(4)"
   TextField "Text field_36" at 564,224 size 204x24; Text 'Step 2'
      Visibility <- "DB_HMI_ARG1_Seq1_S12(4)"
   TextField "Text field_37" at 564,248 size 204x24; Text 'Step 3'
      Visibility <- "DB_HMI_ARG1_Seq1_S13(4)"
   TextField "Text field_38" at 564,272 size 204x24; Text 'Step 4'
      Visibility <- "DB_HMI_ARG1_Seq1_S14(4)"
   TextField "Text field_39" at 564,296 size 204x24; Text 'Step 5'
      Visibility <- "DB_HMI_ARG1_Seq1_S15(4)"
   TextField "Text field_40" at 564,320 size 204x24; Text 'Step 6'
      Visibility <- "DB_HMI_ARG1_Seq1_S16(4)"
   TextField "Text field_41" at 564,344 size 204x24; Text 'Step 7'
      Visibility <- "DB_HMI_ARG1_Seq1_S17(4)"
   TextField "Text field_42" at 564,368 size 204x24; Text 'Step 8'
      Visibility <- "DB_HMI_ARG1_Seq1_S18(4)"
   TextField "Text field_43" at 564,392 size 204x24; Text 'Step 9'
      Visibility <- "DB_HMI_ARG1_Seq1_S19(4)"
   TextField "Text field_44" at 344,138 size 204x24; Text 'Step 0'
      Visibility <- "DB_HMI_ARG1_Seq1_S1(4)"
   TextField "Busy" at 14,134 size 41x22; Text 'Busy'
      Visibility <- "DB_HMI_ARG1_Seq1_Status_Busy(4)"
   TextField "Idle" at 14,134 size 35x22; Text 'Idle'
      Visibility <- "DB_HMI_ARG1_Seq1_Status_Idle(4)"
   Rectangle "rectState" at 0,48 size 56x38
      Appearance <- "CurrentMachineState"
   Button "btnState" at 201,53 size 34x31; TextOff '...'; PictureOff "More_Icon"
      on Click: ActivateScreen("35_Mode_Station_5", 0)
   TextField "Auto" at 67,63 size 35x20; Text 'Auto'
      Visibility <- "DB_HMI_ARG1_Seq1_Status_Auto(4)"
   TextField "Manual" at 69,63 size 34x20; Text 'Man'
      Visibility <- "DB_HMI_ARG1_Seq1_Status_Man(4)"
   TextField "txtStateHeadline" at 65,48 size 123x23; Text 'Mode / Status'

screen "31_Mode_Station_1" 800x480
   Button "Button_5" at 299,208 size 88x48; TextOff 'Stop / AUTO'
      on Press: SetTag("DB_HMI_ARG1_Seq1_Cmd_Auto", 1)
      on Release: SetTag("DB_HMI_ARG1_Seq1_Cmd_Auto", 0)
   Button "Button_6" at 405,208 size 88x48; TextOff 'Reset / MAN'
      on Press: SetTag("DB_HMI_ARG1_Seq1_Cmd_Man", 1)
      on Release: SetTag("DB_HMI_ARG1_Seq1_Cmd_Man", 0)
   Button "Button_1" at 177,283 size 440x40; TextOn 'CLOSE / SCHLIESSEN'; TextOff 'CLOSE / SCHLIESSEN'
      on Click: function_efd93a16()
      Appearance <- "ButtonDown"
   TextField "txtTitleBar" at 16,8 size 495x32; Text 'Operating Mode / Betriebsmodus'
   TextField "txtParameter7_3" at 193,122 size 163x24; Text 'Current Mode / Aktueller Modus'
   TextField "Auto" at 193,149 size 37x20; Text 'Auto'
      Visibility <- "DB_HMI_ARG1_Seq1_Status_Auto"
   TextField "Manual" at 193,149 size 32x20; Text 'Man'
      Visibility <- "DB_HMI_ARG1_Seq1_Status_Man"

screen "32_Mode_Station_2" 800x480
   Button "Button_5" at 299,208 size 88x48; TextOff 'Stop / AUTO'
      on Press: SetTag("DB_HMI_ARG1_Seq1_Cmd_Auto(1)", 1)
      on Release: SetTag("DB_HMI_ARG1_Seq1_Cmd_Auto(1)", 0)
   Button "Button_6" at 405,208 size 88x48; TextOff 'Reset / MAN'
      on Press: SetTag("DB_HMI_ARG1_Seq1_Cmd_Man(1)", 1)
      on Release: SetTag("DB_HMI_ARG1_Seq1_Cmd_Man(1)", 0)
   Button "Button_1" at 177,283 size 440x40; TextOn 'CLOSE / SCHLIESSEN'; TextOff 'CLOSE / SCHLIESSEN'
      on Click: function_efd93a16()
      Appearance <- "ButtonDown"
   TextField "txtTitleBar" at 16,8 size 495x32; Text 'Operating Mode / Betriebsmodus'
   TextField "txtParameter7_3" at 193,122 size 163x24; Text 'Current Mode / Aktueller Modus'
   TextField "Auto" at 193,149 size 37x20; Text 'Auto'
      Visibility <- "DB_HMI_ARG1_Seq1_Status_Auto(1)"
   TextField "Manual" at 193,148 size 32x20; Text 'Man'
      Visibility <- "DB_HMI_ARG1_Seq1_Status_Man(1)"